       "DB_CrossCut_1_HMI".tHMR.xManualCommandEnabled := "FB_CrossCuts_1_V1_00_IDB".tHMR.xManComEn;
       "DB_CrossCut_1_HMI".tHMR.tManCmd.xManJogFwdFdbk := "FB_CrossCuts_1_V1_00_IDB".tHMR.tManCmd.xManJogFwdFdbk;
       "DB_CrossCut_1_HMI".tHMR.tManCmd.xManJogBckFdbk := "FB_CrossCuts_1_V1_00_IDB".tHMR.tManCmd.xManJogBckFdbk;
       "DB_CrossCut_1_HMI".tHMR.tManCmd.xManCarriageDownFdbk := "FB_CrossCuts_1_V1_00_IDB".tHMR.tManCmd.xManCarriageDownFdbk;
       "DB_CrossCut_1_HMI".tHMR.tManCmd.xManFireONFdbk := "FB_CrossCuts_1_V1_00_IDB".tHMR.tManCmd.xManFireONFdbk;
       "DB_CrossCut_1_HMI".tHMR.tManCmd.xManOilONFdbk := "FB_CrossCuts_1_V1_00_IDB".tHMR.tManCmd.xManOilONFdbk;

       "DB_CrossCut_1_HMI".tHMR.dDistanceSnaproll_cmm := "FB_CrossCuts_1_V1_00_IDB".tHMR.dDistanceFromSnaproll_cmm;
       "DB_CrossCut_1_HMI".tHMR.dStatus := "FB_CrossCuts_1_V1_00_IDB".tHMR.dStatus;
       "DB_CrossCut_1_HMI".tHMR.dXCutActualStatus := "FB_CrossCuts_1_V1_00_IDB".tHMR.dXCutActualStatus;
       "DB_CrossCut_1_HMI".tHMR.dXCutStatusRequest:="FB_CrossCuts_1_V1_00_IDB".tHMR.dXCutStatusRequest;
       "DB_CrossCut_1_HMI".tHMR.dDistanceFromCenterLine_cmm := "FB_CrossCuts_1_V1_00_IDB".tHMR.dDistanceFromCenterLine_cmm;
       "DB_CrossCut_1_HMI".tHMR.dAngleValue_uDegree := "FB_CrossCuts_1_V1_00_IDB".tHMR.dAngleValue_uDegree;
       "DB_CrossCut_1_HMI".tHMR.dActualCutPosRequest := "FB_CrossCuts_1_V1_00_IDB".tHMR.dActualCutPosRequest;
       "DB_CrossCut_1_HMI".tHMR.dCarriagePosition_cmm := "FB_CrossCuts_1_V1_00_IDB".tHMR.dCarriagePosition_cmm;

       "DB_CrossCut_1_HMI".tHMR.rHeadUsage_km := "FB_CrossCuts_1_V1_00_IDB".tHMR.rHeadUsage_km;

       //Move CROSS CUT #1 HMW 
       "FB_CrossCuts_1_V1_00_IDB".tHMW.xCutBreakEnabled := "DB_CrossCut_1_HMI".tHMW.xCutBreakEnabled;
       "FB_CrossCuts_1_V1_00_IDB".tHMW.xUpdateDistSnap := "DB_CrossCut_1_HMI".tHMW.xUpdateDistanceSnaproll;
       "FB_CrossCuts_1_V1_00_IDB".tHMW.xUpdateAngleValue := "DB_CrossCut_1_HMI".tHMW.xUpdateAngleValue;
       "FB_CrossCuts_1_V1_00_IDB".tHMW.xIncAngleValue := "DB_CrossCut_1_HMI".tHMW.xIncAngleValue;
       "FB_CrossCuts_1_V1_00_IDB".tHMW.xDecAngleValue := "DB_CrossCut_1_HMI".tHMW.xDecAngleValue;
       "FB_CrossCuts_1_V1_00_IDB".tHMW.xUpdateDistCenterLine := "DB_CrossCut_1_HMI".tHMW.xUpdateDistCenterLine;
       "FB_CrossCuts_1_V1_00_IDB".tHMW.xCalibDistRequest := "DB_CrossCut_1_HMI".tHMW.xCalibDistRequest;
       "FB_CrossCuts_1_V1_00_IDB".tHMW.xCalibDiagRequest := "DB_CrossCut_1_HMI".tHMW.xCalibDiagRequest;
       "FB_CrossCuts_1_V1_00_IDB".tHMW.xCutOperator := "DB_CrossCut_1_HMI".tHMW.xCutOperator;
       "FB_CrossCuts_1_V1_00_IDB".tHMW.xCutGross := "DB_CrossCut_1_HMI".tHMW.xCutGross;
       "FB_CrossCuts_1_V1_00_IDB".tHMW.xCutNet := "DB_CrossCut_1_HMI".tHMW.xCutNet;
       "FB_CrossCuts_1_V1_00_IDB".tHMW.xCutYCut := "DB_CrossCut_1_HMI".tHMW.xCutYCut;
       "FB_CrossCuts_1_V1_00_IDB".tHMW.xEnDisManCom := "DB_CrossCut_1_HMI".tHMW.xEnableManualCommand;
       "FB_CrossCuts_1_V1_00_IDB".tHMW.xResetHeadUsage := "DB_CrossCut_1_HMI".tHMW.xResetHeadUsage;

       "FB_CrossCuts_1_V1_00_IDB".tHMW.tManCmd.xMan_JogForward := "DB_CrossCut_1_HMI".tHMW.tManCmd.xMan_JogForward;
       "FB_CrossCuts_1_V1_00_IDB".tHMW.tManCmd.xMan_JobBackward := "DB_CrossCut_1_HMI".tHMW.tManCmd.xMan_JobBackward;
       "FB_CrossCuts_1_V1_00_IDB".tHMW.tManCmd.xMan_CarriageDown := "DB_CrossCut_1_HMI".tHMW.tManCmd.xMan_CarriageDown;
       "FB_CrossCuts_1_V1_00_IDB".tHMW.tManCmd.xMan_FireOn := "DB_CrossCut_1_HMI".tHMW.tManCmd.xMan_FireOn;
       "FB_CrossCuts_1_V1_00_IDB".tHMW.tManCmd.xMan_OilOn := "DB_CrossCut_1_HMI".tHMW.tManCmd.xMan_OilOn;



      "FB_CrossCuts_1_V1_00_IDB".tHMW.dOperStartCutPos_cmm := "DB_CrossCut_1_HMI".tHMW.dOperStartCutPos_cmm;
      "FB_CrossCuts_1_V1_00_IDB".tHMW.dOperEndCutPos_cmm := "DB_CrossCut_1_HMI".tHMW.dOperEndCutPos_cmm;
      "FB_CrossCuts_1_V1_00_IDB".tHMW.dDescReactTime_ms := "DB_CrossCut_1_HMI".tHMW.dDescReactTime_ms;
      "FB_CrossCuts_1_V1_00_IDB".tHMW.dRaiseReactTime_ms := "DB_CrossCut_1_HMI".tHMW.dRaiseReactTime_ms;

      "FB_CrossCuts_1_V1_00_IDB".tHMW.dFireONReactTime_ms := "DB_CrossCut_1_HMI".tHMW.dFireONReactTime_ms;
      "FB_CrossCuts_1_V1_00_IDB".tHMW.dFireOFFReactTime_ms := "DB_CrossCut_1_HMI".tHMW.dFireOFFReactTime_ms;
      "FB_CrossCuts_1_V1_00_IDB".tHMW.dOilONDelay_ms := "DB_CrossCut_1_HMI".tHMW.dOilONDelay_ms;
      "FB_CrossCuts_1_V1_00_IDB".tHMW.dOilOFFDelay_ms := "DB_CrossCut_1_HMI".tHMW.dOilOFFDelay_ms;

      "FB_CrossCuts_1_V1_00_IDB".tHMW.dCutStartOffsetDelay_cmm := "DB_CrossCut_1_HMI".tHMW.dCutStartOffsetDelay_cmm;
      "FB_CrossCuts_1_V1_00_IDB".tHMW.dCutEndOffsetDelay_cmm := "DB_CrossCut_1_HMI".tHMW.dCutEndOffsetDelay_cmm;

      "FB_CrossCuts_1_V1_00_IDB".tHMW.dDistanceFromSnaproll_cmm := "DB_CrossCut_1_HMI".tHMW.dDistanceSnaproll_cmm;
      "FB_CrossCuts_1_V1_00_IDB".tHMW.dAngleValue_uDegree := "DB_CrossCut_1_HMI".tHMW.dAngleValue_uDegree;
      "FB_CrossCuts_1_V1_00_IDB".tHMW.dDistanceFromCenterLine_cmm := "DB_CrossCut_1_HMI".tHMW.dDistanceFromCenterLine_cmm;
      "FB_CrossCuts_1_V1_00_IDB".tHMW.dDistTeoLength_cmm := "DB_CrossCut_1_HMI".tHMW.dDistTeoLength_cmm;
      "FB_CrossCuts_1_V1_00_IDB".tHMW.dDistRealLength_cmm := "DB_CrossCut_1_HMI".tHMW.dDistRealLength_cmm;

      "FB_CrossCuts_1_V1_00_IDB".tHMW.dDiagRealWidth_cmm := "DB_CrossCut_1_HMI".tHMW.dDiagRealWidth_cmm;
       "FB_CrossCuts_1_V1_00_IDB".tHMW.dDiagRealLength_cmm := "DB_CrossCut_1_HMI".tHMW.dDiagRealLength_cmm;
       "FB_CrossCuts_1_V1_00_IDB".tHMW.dDiagGlassFlow_cmm := "DB_CrossCut_1_HMI".tHMW.dDiagGlassFlow_cmm;
       "FB_CrossCuts_1_V1_00_IDB".tHMW.dDiagGlassOppFlow_cmm := "DB_CrossCut_1_HMI".tHMW.dDiagGlassOppFlow_cmm;

       "FB_CrossCuts_1_V1_00_IDB".tHMW.dCuttingPressure_mN := "DB_CrossCut_1_HMI".tHMW.dCuttingPressure_mN;
       "FB_CrossCuts_1_V1_00_IDB".tHMW.dPosOffset_cmm := "DB_CrossCut_1_HMI".tHMW.dPosOffset_cmm;

       "FB_CrossCuts_1_V1_00_IDB".tHMW.dCutPriority := "DB_CrossCut_1_HMI".tHMW.dCutPriority;

       //Move CROSS CUT #1 ALM
       "DB_CrossCut_1_HMI".tALM := "FB_CrossCuts_1_V1_00_IDB".tALM;



       //Move CROSS CUT #2 HMR 

       "DB_CrossCut_2_HMI".tHMR.xManualCommandEnabled := "FB_CrossCuts_2_V1_00_IDB".tHMR.xManComEn;
       "DB_CrossCut_2_HMI".tHMR.tManCmd.xManJogFwdFdbk := "FB_CrossCuts_2_V1_00_IDB".tHMR.tManCmd.xManJogFwdFdbk;
       "DB_CrossCut_2_HMI".tHMR.tManCmd.xManJogBckFdbk := "FB_CrossCuts_2_V1_00_IDB".tHMR.tManCmd.xManJogBckFdbk;
       "DB_CrossCut_2_HMI".tHMR.tManCmd.xManCarriageDownFdbk := "FB_CrossCuts_2_V1_00_IDB".tHMR.tManCmd.xManCarriageDownFdbk;
       "DB_CrossCut_2_HMI".tHMR.tManCmd.xManFireONFdbk := "FB_CrossCuts_2_V1_00_IDB".tHMR.tManCmd.xManFireONFdbk;
       "DB_CrossCut_2_HMI".tHMR.tManCmd.xManOilONFdbk := "FB_CrossCuts_2_V1_00_IDB".tHMR.tManCmd.xManOilONFdbk;

       "DB_CrossCut_2_HMI".tHMR.dDistanceSnaproll_cmm := "FB_CrossCuts_2_V1_00_IDB".tHMR.dDistanceFromSnaproll_cmm;
       "DB_CrossCut_2_HMI".tHMR.dStatus := "FB_CrossCuts_2_V1_00_IDB".tHMR.dStatus;
       "DB_CrossCut_2_HMI".tHMR.dXCutActualStatus := "FB_CrossCuts_2_V1_00_IDB".tHMR.dXCutActualStatus;
       "DB_CrossCut_2_HMI".tHMR.dXCutStatusRequest := "FB_CrossCuts_2_V1_00_IDB".tHMR.dXCutStatusRequest;
       "DB_CrossCut_2_HMI".tHMR.dDistanceFromCenterLine_cmm := "FB_CrossCuts_2_V1_00_IDB".tHMR.dDistanceFromCenterLine_cmm;
       "DB_CrossCut_2_HMI".tHMR.dAngleValue_uDegree := "FB_CrossCuts_2_V1_00_IDB".tHMR.dAngleValue_uDegree;
       "DB_CrossCut_2_HMI".tHMR.dActualCutPosRequest := "FB_CrossCuts_2_V1_00_IDB".tHMR.dActualCutPosRequest;
       "DB_CrossCut_2_HMI".tHMR.dCarriagePosition_cmm := "FB_CrossCuts_2_V1_00_IDB".tHMR.dCarriagePosition_cmm;

       "DB_CrossCut_2_HMI".tHMR.rHeadUsage_km := "FB_CrossCuts_2_V1_00_IDB".tHMR.rHeadUsage_km;

       //Move CROSS CUT #2 HMW 
       "FB_CrossCuts_2_V1_00_IDB".tHMW.xCutBreakEnabled := "DB_CrossCut_2_HMI".tHMW.xCutBreakEnabled;
       "FB_CrossCuts_2_V1_00_IDB".tHMW.xUpdateDistSnap := "DB_CrossCut_2_HMI".tHMW.xUpdateDistanceSnaproll;
       "FB_CrossCuts_2_V1_00_IDB".tHMW.xUpdateAngleValue := "DB_CrossCut_2_HMI".tHMW.xUpdateAngleValue;
       "FB_CrossCuts_2_V1_00_IDB".tHMW.xIncAngleValue := "DB_CrossCut_2_HMI".tHMW.xIncAngleValue;
       "FB_CrossCuts_2_V1_00_IDB".tHMW.xDecAngleValue := "DB_CrossCut_2_HMI".tHMW.xDecAngleValue;
       "FB_CrossCuts_2_V1_00_IDB".tHMW.xUpdateDistCenterLine := "DB_CrossCut_2_HMI".tHMW.xUpdateDistCenterLine;
       "FB_CrossCuts_2_V1_00_IDB".tHMW.xCalibDistRequest := "DB_CrossCut_2_HMI".tHMW.xCalibDistRequest;
       "FB_CrossCuts_2_V1_00_IDB".tHMW.xCalibDiagRequest := "DB_CrossCut_2_HMI".tHMW.xCalibDiagRequest;
       "FB_CrossCuts_2_V1_00_IDB".tHMW.xCutOperator := "DB_CrossCut_2_HMI".tHMW.xCutOperator;
       "FB_CrossCuts_2_V1_00_IDB".tHMW.xCutGross := "DB_CrossCut_2_HMI".tHMW.xCutGross;
       "FB_CrossCuts_2_V1_00_IDB".tHMW.xCutNet := "DB_CrossCut_2_HMI".tHMW.xCutNet;
       "FB_CrossCuts_2_V1_00_IDB".tHMW.xCutYCut := "DB_CrossCut_2_HMI".tHMW.xCutYCut;
       "FB_CrossCuts_2_V1_00_IDB".tHMW.xEnDisManCom := "DB_CrossCut_2_HMI".tHMW.xEnableManualCommand;
       "FB_CrossCuts_2_V1_00_IDB".tHMW.xResetHeadUsage := "DB_CrossCut_2_HMI".tHMW.xResetHeadUsage;

       "FB_CrossCuts_2_V1_00_IDB".tHMW.tManCmd.xMan_JogForward := "DB_CrossCut_2_HMI".tHMW.tManCmd.xMan_JogForward;
       "FB_CrossCuts_2_V1_00_IDB".tHMW.tManCmd.xMan_JobBackward := "DB_CrossCut_2_HMI".tHMW.tManCmd.xMan_JobBackward;
       "FB_CrossCuts_2_V1_00_IDB".tHMW.tManCmd.xMan_CarriageDown := "DB_CrossCut_2_HMI".tHMW.tManCmd.xMan_CarriageDown;
       "FB_CrossCuts_2_V1_00_IDB".tHMW.tManCmd.xMan_FireOn := "DB_CrossCut_2_HMI".tHMW.tManCmd.xMan_FireOn;
       "FB_CrossCuts_2_V1_00_IDB".tHMW.tManCmd.xMan_OilOn := "DB_CrossCut_2_HMI".tHMW.tManCmd.xMan_OilOn;



       "FB_CrossCuts_2_V1_00_IDB".tHMW.dOperStartCutPos_cmm := "DB_CrossCut_2_HMI".tHMW.dOperStartCutPos_cmm;
       "FB_CrossCuts_2_V1_00_IDB".tHMW.dOperEndCutPos_cmm := "DB_CrossCut_2_HMI".tHMW.dOperEndCutPos_cmm;
       "FB_CrossCuts_2_V1_00_IDB".tHMW.dDescReactTime_ms := "DB_CrossCut_2_HMI".tHMW.dDescReactTime_ms;
       "FB_CrossCuts_2_V1_00_IDB".tHMW.dRaiseReactTime_ms := "DB_CrossCut_2_HMI".tHMW.dRaiseReactTime_ms;

       "FB_CrossCuts_2_V1_00_IDB".tHMW.dFireONReactTime_ms := "DB_CrossCut_2_HMI".tHMW.dFireONReactTime_ms;
       "FB_CrossCuts_2_V1_00_IDB".tHMW.dFireOFFReactTime_ms := "DB_CrossCut_2_HMI".tHMW.dFireOFFReactTime_ms;
       "FB_CrossCuts_2_V1_00_IDB".tHMW.dOilONDelay_ms := "DB_CrossCut_2_HMI".tHMW.dOilONDelay_ms;
       "FB_CrossCuts_2_V1_00_IDB".tHMW.dOilOFFDelay_ms := "DB_CrossCut_2_HMI".tHMW.dOilOFFDelay_ms;

       "FB_CrossCuts_2_V1_00_IDB".tHMW.dCutStartOffsetDelay_cmm := "DB_CrossCut_2_HMI".tHMW.dCutStartOffsetDelay_cmm;
       "FB_CrossCuts_2_V1_00_IDB".tHMW.dCutEndOffsetDelay_cmm := "DB_CrossCut_2_HMI".tHMW.dCutEndOffsetDelay_cmm;

       "FB_CrossCuts_2_V1_00_IDB".tHMW.dDistanceFromSnaproll_cmm := "DB_CrossCut_2_HMI".tHMW.dDistanceSnaproll_cmm;
       "FB_CrossCuts_2_V1_00_IDB".tHMW.dAngleValue_uDegree := "DB_CrossCut_2_HMI".tHMW.dAngleValue_uDegree;
       "FB_CrossCuts_2_V1_00_IDB".tHMW.dDistanceFromCenterLine_cmm := "DB_CrossCut_2_HMI".tHMW.dDistanceFromCenterLine_cmm;
       "FB_CrossCuts_2_V1_00_IDB".tHMW.dDistTeoLength_cmm := "DB_CrossCut_2_HMI".tHMW.dDistTeoLength_cmm;
       "FB_CrossCuts_2_V1_00_IDB".tHMW.dDistRealLength_cmm := "DB_CrossCut_2_HMI".tHMW.dDistRealLength_cmm;

       "FB_CrossCuts_2_V1_00_IDB".tHMW.dDiagRealWidth_cmm := "DB_CrossCut_2_HMI".tHMW.dDiagRealWidth_cmm;
       "FB_CrossCuts_2_V1_00_IDB".tHMW.dDiagRealLength_cmm := "DB_CrossCut_2_HMI".tHMW.dDiagRealLength_cmm;
       "FB_CrossCuts_2_V1_00_IDB".tHMW.dDiagGlassFlow_cmm := "DB_CrossCut_2_HMI".tHMW.dDiagGlassFlow_cmm;
       "FB_CrossCuts_2_V1_00_IDB".tHMW.dDiagGlassOppFlow_cmm := "DB_CrossCut_2_HMI".tHMW.dDiagGlassOppFlow_cmm;

       "FB_CrossCuts_2_V1_00_IDB".tHMW.dCuttingPressure_mN := "DB_CrossCut_2_HMI".tHMW.dCuttingPressure_mN;
       "FB_CrossCuts_2_V1_00_IDB".tHMW.dPosOffset_cmm := "DB_CrossCut_2_HMI".tHMW.dPosOffset_cmm;

       "FB_CrossCuts_2_V1_00_IDB".tHMW.dCutPriority := "DB_CrossCut_2_HMI".tHMW.dCutPriority;

       //Move CROSS CUT #2 ALM
       "DB_CrossCut_2_HMI".tALM := "FB_CrossCuts_2_V1_00_IDB".tALM;



       //Move CROSS CUT #3 HMR 

       "DB_CrossCut_3_HMI".tHMR.xManualCommandEnabled := "FB_CrossCuts_3_V1_00_IDB".tHMR.xManComEn;
       "DB_CrossCut_3_HMI".tHMR.tManCmd.xManJogFwdFdbk := "FB_CrossCuts_3_V1_00_IDB".tHMR.tManCmd.xManJogFwdFdbk;
       "DB_CrossCut_3_HMI".tHMR.tManCmd.xManJogBckFdbk := "FB_CrossCuts_3_V1_00_IDB".tHMR.tManCmd.xManJogBckFdbk;
       "DB_CrossCut_3_HMI".tHMR.tManCmd.xManCarriageDownFdbk := "FB_CrossCuts_3_V1_00_IDB".tHMR.tManCmd.xManCarriageDownFdbk;
       "DB_CrossCut_3_HMI".tHMR.tManCmd.xManFireONFdbk := "FB_CrossCuts_3_V1_00_IDB".tHMR.tManCmd.xManFireONFdbk;
       "DB_CrossCut_3_HMI".tHMR.tManCmd.xManOilONFdbk := "FB_CrossCuts_3_V1_00_IDB".tHMR.tManCmd.xManOilONFdbk;

       "DB_CrossCut_3_HMI".tHMR.dDistanceSnaproll_cmm := "FB_CrossCuts_3_V1_00_IDB".tHMR.dDistanceFromSnaproll_cmm;
       "DB_CrossCut_3_HMI".tHMR.dStatus := "FB_CrossCuts_3_V1_00_IDB".tHMR.dStatus;
       "DB_CrossCut_3_HMI".tHMR.dXCutActualStatus := "FB_CrossCuts_3_V1_00_IDB".tHMR.dXCutActualStatus;
       "DB_CrossCut_3_HMI".tHMR.dXCutStatusRequest := "FB_CrossCuts_3_V1_00_IDB".tHMR.dXCutStatusRequest;
       "DB_CrossCut_3_HMI".tHMR.dDistanceFromCenterLine_cmm := "FB_CrossCuts_3_V1_00_IDB".tHMR.dDistanceFromCenterLine_cmm;
       "DB_CrossCut_3_HMI".tHMR.dAngleValue_uDegree := "FB_CrossCuts_3_V1_00_IDB".tHMR.dAngleValue_uDegree;
       "DB_CrossCut_3_HMI".tHMR.dActualCutPosRequest := "FB_CrossCuts_3_V1_00_IDB".tHMR.dActualCutPosRequest;
       "DB_CrossCut_3_HMI".tHMR.dCarriagePosition_cmm := "FB_CrossCuts_3_V1_00_IDB".tHMR.dCarriagePosition_cmm;

       "DB_CrossCut_3_HMI".tHMR.rHeadUsage_km := "FB_CrossCuts_3_V1_00_IDB".tHMR.rHeadUsage_km;

       //Move CROSS CUT #3 HMW 
       "FB_CrossCuts_3_V1_00_IDB".tHMW.xCutBreakEnabled := "DB_CrossCut_3_HMI".tHMW.xCutBreakEnabled;
       "FB_CrossCuts_3_V1_00_IDB".tHMW.xUpdateDistSnap := "DB_CrossCut_3_HMI".tHMW.xUpdateDistanceSnaproll;
       "FB_CrossCuts_3_V1_00_IDB".tHMW.xUpdateAngleValue := "DB_CrossCut_3_HMI".tHMW.xUpdateAngleValue;
       "FB_CrossCuts_3_V1_00_IDB".tHMW.xIncAngleValue := "DB_CrossCut_3_HMI".tHMW.xIncAngleValue;
       "FB_CrossCuts_3_V1_00_IDB".tHMW.xDecAngleValue := "DB_CrossCut_3_HMI".tHMW.xDecAngleValue;
       "FB_CrossCuts_3_V1_00_IDB".tHMW.xUpdateDistCenterLine := "DB_CrossCut_3_HMI".tHMW.xUpdateDistCenterLine;
       "FB_CrossCuts_3_V1_00_IDB".tHMW.xCalibDistRequest := "DB_CrossCut_3_HMI".tHMW.xCalibDistRequest;
       "FB_CrossCuts_3_V1_00_IDB".tHMW.xCalibDiagRequest := "DB_CrossCut_3_HMI".tHMW.xCalibDiagRequest;
       "FB_CrossCuts_3_V1_00_IDB".tHMW.xCutOperator := "DB_CrossCut_3_HMI".tHMW.xCutOperator;
       "FB_CrossCuts_3_V1_00_IDB".tHMW.xCutGross := "DB_CrossCut_3_HMI".tHMW.xCutGross;
       "FB_CrossCuts_3_V1_00_IDB".tHMW.xCutNet := "DB_CrossCut_3_HMI".tHMW.xCutNet;
       "FB_CrossCuts_3_V1_00_IDB".tHMW.xCutYCut := "DB_CrossCut_3_HMI".tHMW.xCutYCut;
       "FB_CrossCuts_3_V1_00_IDB".tHMW.xEnDisManCom := "DB_CrossCut_3_HMI".tHMW.xEnableManualCommand;
       "FB_CrossCuts_3_V1_00_IDB".tHMW.xResetHeadUsage := "DB_CrossCut_3_HMI".tHMW.xResetHeadUsage;

       "FB_CrossCuts_3_V1_00_IDB".tHMW.tManCmd.xMan_JogForward := "DB_CrossCut_3_HMI".tHMW.tManCmd.xMan_JogForward;
       "FB_CrossCuts_3_V1_00_IDB".tHMW.tManCmd.xMan_JobBackward := "DB_CrossCut_3_HMI".tHMW.tManCmd.xMan_JobBackward;
       "FB_CrossCuts_3_V1_00_IDB".tHMW.tManCmd.xMan_CarriageDown := "DB_CrossCut_3_HMI".tHMW.tManCmd.xMan_CarriageDown;
       "FB_CrossCuts_3_V1_00_IDB".tHMW.tManCmd.xMan_FireOn := "DB_CrossCut_3_HMI".tHMW.tManCmd.xMan_FireOn;
       "FB_CrossCuts_3_V1_00_IDB".tHMW.tManCmd.xMan_OilOn := "DB_CrossCut_3_HMI".tHMW.tManCmd.xMan_OilOn;



       "FB_CrossCuts_3_V1_00_IDB".tHMW.dOperStartCutPos_cmm := "DB_CrossCut_3_HMI".tHMW.dOperStartCutPos_cmm;
       "FB_CrossCuts_3_V1_00_IDB".tHMW.dOperEndCutPos_cmm := "DB_CrossCut_3_HMI".tHMW.dOperEndCutPos_cmm;
       "FB_CrossCuts_3_V1_00_IDB".tHMW.dDescReactTime_ms := "DB_CrossCut_3_HMI".tHMW.dDescReactTime_ms;
       "FB_CrossCuts_3_V1_00_IDB".tHMW.dRaiseReactTime_ms := "DB_CrossCut_3_HMI".tHMW.dRaiseReactTime_ms;

       "FB_CrossCuts_3_V1_00_IDB".tHMW.dFireONReactTime_ms := "DB_CrossCut_3_HMI".tHMW.dFireONReactTime_ms;
       "FB_CrossCuts_3_V1_00_IDB".tHMW.dFireOFFReactTime_ms := "DB_CrossCut_3_HMI".tHMW.dFireOFFReactTime_ms;
       "FB_CrossCuts_3_V1_00_IDB".tHMW.dOilONDelay_ms := "DB_CrossCut_3_HMI".tHMW.dOilONDelay_ms;
       "FB_CrossCuts_3_V1_00_IDB".tHMW.dOilOFFDelay_ms := "DB_CrossCut_3_HMI".tHMW.dOilOFFDelay_ms;

       "FB_CrossCuts_3_V1_00_IDB".tHMW.dCutStartOffsetDelay_cmm := "DB_CrossCut_3_HMI".tHMW.dCutStartOffsetDelay_cmm;
       "FB_CrossCuts_3_V1_00_IDB".tHMW.dCutEndOffsetDelay_cmm := "DB_CrossCut_3_HMI".tHMW.dCutEndOffsetDelay_cmm;

       "FB_CrossCuts_3_V1_00_IDB".tHMW.dDistanceFromSnaproll_cmm := "DB_CrossCut_3_HMI".tHMW.dDistanceSnaproll_cmm;
       "FB_CrossCuts_3_V1_00_IDB".tHMW.dAngleValue_uDegree := "DB_CrossCut_3_HMI".tHMW.dAngleValue_uDegree;
       "FB_CrossCuts_3_V1_00_IDB".tHMW.dDistanceFromCenterLine_cmm := "DB_CrossCut_3_HMI".tHMW.dDistanceFromCenterLine_cmm;
       "FB_CrossCuts_3_V1_00_IDB".tHMW.dDistTeoLength_cmm := "DB_CrossCut_3_HMI".tHMW.dDistTeoLength_cmm;
       "FB_CrossCuts_3_V1_00_IDB".tHMW.dDistRealLength_cmm := "DB_CrossCut_3_HMI".tHMW.dDistRealLength_cmm;

       "FB_CrossCuts_3_V1_00_IDB".tHMW.dDiagRealWidth_cmm := "DB_CrossCut_3_HMI".tHMW.dDiagRealWidth_cmm;
       "FB_CrossCuts_3_V1_00_IDB".tHMW.dDiagRealLength_cmm := "DB_CrossCut_3_HMI".tHMW.dDiagRealLength_cmm;
       "FB_CrossCuts_3_V1_00_IDB".tHMW.dDiagGlassFlow_cmm := "DB_CrossCut_3_HMI".tHMW.dDiagGlassFlow_cmm;
       "FB_CrossCuts_3_V1_00_IDB".tHMW.dDiagGlassOppFlow_cmm := "DB_CrossCut_3_HMI".tHMW.dDiagGlassOppFlow_cmm;

       "FB_CrossCuts_3_V1_00_IDB".tHMW.dCuttingPressure_mN := "DB_CrossCut_3_HMI".tHMW.dCuttingPressure_mN;
       "FB_CrossCuts_3_V1_00_IDB".tHMW.dPosOffset_cmm := "DB_CrossCut_3_HMI".tHMW.dPosOffset_cmm;

       "FB_CrossCuts_3_V1_00_IDB".tHMW.dCutPriority := "DB_CrossCut_3_HMI".tHMW.dCutPriority;

       //Move CROSS CUT #3 ALM
       "DB_CrossCut_3_HMI".tALM := "FB_CrossCuts_3_V1_00_IDB".tALM;



       //Move YCUT 1 HMR
       "DB_YCut_1_HMI".tHMR.dDistanceSnaproll_cmm := "FB_YCuts1_V1_00_IDB".tHMR.dDistanceFromSnaproll_cmm;
       //Move YCUT 1  HMW
       "FB_YCuts1_V1_00_IDB".tHMW.xUpdateDistSnap := "DB_YCut_1_HMI".tHMW.xUpdateDistanceSnaproll;
       "FB_YCuts1_V1_00_IDB".tHMW.dDistanceFromSnaproll_cmm := "DB_YCut_1_HMI".tHMW.dDistanceSnaproll_cmm;
       //Move YCUT 1  ALM 
       "DB_YCut_1_HMI".tALM.tF := "FB_YCuts1_V1_00_IDB".tALM.tF;
       "DB_YCut_1_HMI".tALM.tS := "FB_YCuts1_V1_00_IDB".tALM.tS;
       "DB_YCut_1_HMI".tALM.tW:= "FB_YCuts1_V1_00_IDB".tALM.tW;

       //Move YCUT 2 HMR
       "DB_YCut_2_HMI".tHMR.dDistanceSnaproll_cmm := "FB_YCuts2_V1_00_IDB".tHMR.dDistanceFromSnaproll_cmm;
       //Move YCUT 2  HMW
       "FB_YCuts2_V1_00_IDB".tHMW.xUpdateDistSnap := "DB_YCut_2_HMI".tHMW.xUpdateDistanceSnaproll;
       "FB_YCuts2_V1_00_IDB".tHMW.dDistanceFromSnaproll_cmm := "DB_YCut_2_HMI".tHMW.dDistanceSnaproll_cmm;
       //Move YCUT 1  ALM 
       "DB_YCut_2_HMI".tALM.tF := "FB_YCuts2_V1_00_IDB".tALM.tF;
       "DB_YCut_2_HMI".tALM.tS := "FB_YCuts2_V1_00_IDB".tALM.tS;
       "DB_YCut_2_HMI".tALM.tW := "FB_YCuts2_V1_00_IDB".tALM.tW;

       //Move Marker M220 HMR
       "DB_Marker_HMI".tHMR.dSpare0 :="FB_Markers_V1.00_IDB".tHMR.dSpare;
       //Move Marker M220  HMW
       "FB_Markers_V1.00_IDB".tHMW.dSpare :=  "DB_Marker_HMI".tHMW.dSpare0;
       //Move Marker M220 ALM  
       "DB_Marker_HMI".tALM.tF := "FB_Markers_V1.00_IDB".tALM.tF;
       "DB_Marker_HMI".tALM.tS := "FB_Markers_V1.00_IDB".tALM.tS;
       "DB_Marker_HMI".tALM.tW := "FB_Markers_V1.00_IDB".tALM.tW;

       //Move DIGITIZER #1 HMR
       "DB_Digitizer_1_HMI".tHMR.xManualCommandEnabled := "FB_Digitizer_1_V1_00_IDB".tHMR.xManComEn;
       "DB_Digitizer_1_HMI".tHMR.tManCmd.xMan_DescEncFdbk:= "FB_Digitizer_1_V1_00_IDB".tHMR.xMan_DescEncFdbk;
       "DB_Digitizer_1_HMI".tHMR.dEncoderStatus := "FB_Digitizer_1_V1_00_IDB".tHMR.dEncoderStatus;
       "DB_Digitizer_1_HMI".tHMR.dFm152Status := "FB_Digitizer_1_V1_00_IDB".tHMR.dFm152Status;
       "DB_Digitizer_1_HMI".tHMR.dActualEncoderSpeed_mm_min := "FB_Digitizer_1_V1_00_IDB".tHMR.dActualEncoderSpeed_mm_min;
       "DB_Digitizer_1_HMI".tHMR.dCalibrationF1Unit_unit := "FB_Digitizer_1_V1_00_IDB".tHMR.dCalibrationF1Unit_unit;
       "DB_Digitizer_1_HMI".tHMR.dCalibrationF2Unit_unit := "FB_Digitizer_1_V1_00_IDB".tHMR.dCalibrationF2Unit_unit;
       "DB_Digitizer_1_HMI".tHMR.dCalibrationCardF1Unit_unit := "FB_Digitizer_1_V1_00_IDB".tHMR.dCalibrationCardF1Unit_unit;
       "DB_Digitizer_1_HMI".tHMR.dCalibrationCardF2Unit_unit := "FB_Digitizer_1_V1_00_IDB".tHMR.dCalibrationCardF2Unit_unit;


       //Move DIGITIZER #1  HMW
       "FB_Digitizer_1_V1_00_IDB".tHMW.xCalibUpdateF1 := "DB_Digitizer_1_HMI".tHMW.xCalibRequest;
       "FB_Digitizer_1_V1_00_IDB".tHMW.xCalibUpdateF2 := "DB_Digitizer_1_HMI".tHMW.xCalibUpdateF1;
       "FB_Digitizer_1_V1_00_IDB".tHMW.xCalibRequest := "DB_Digitizer_1_HMI".tHMW.xCalibUpdateF2;
       "FB_Digitizer_1_V1_00_IDB".tHMW.xMan_DescentEnc:="DB_Digitizer_1_HMI".tHMW.tManCmd.xMan_DescentEnc;
       "FB_Digitizer_1_V1_00_IDB".tHMW.xGlassSensorEnabled := "DB_Digitizer_1_HMI".tHMW.xGlassSensorEnabled;
       "FB_Digitizer_1_V1_00_IDB".tHMW.xEnDisManCom := "DB_Digitizer_1_HMI".tHMW.xEnableManualCommand;
       "FB_Digitizer_1_V1_00_IDB".tHMW.dCalibTheoLength_cmm := "DB_Digitizer_1_HMI".tHMW.dCalibTheoLength_cmm;
       "FB_Digitizer_1_V1_00_IDB".tHMW.dCalibRealLength_cmm := "DB_Digitizer_1_HMI".tHMW.dCalibRealLength_cmm;
       "FB_Digitizer_1_V1_00_IDB".tHMW.dCalibWriteF1_unit := "DB_Digitizer_1_HMI".tHMW.dCalibWriteF1_unit;
       "FB_Digitizer_1_V1_00_IDB".tHMW.dCalibWriteF2_unit := "DB_Digitizer_1_HMI".tHMW.dCalibWriteF2_unit;
       "FB_Digitizer_1_V1_00_IDB".tHMW.dRequestJogSpeed_mm_min := "DB_Digitizer_1_HMI".tHMW.dRequestJogSpeed_mm_min;




       //Move DIGITIZER #1 ALM  
       "DB_Digitizer_1_HMI".tALM.tS := "FB_Digitizer_1_V1_00_IDB".tALM.tS;
       "DB_Digitizer_1_HMI".tALM.tF := "FB_Digitizer_1_V1_00_IDB".tALM.tF;
       "DB_Digitizer_1_HMI".tALM.tW := "FB_Digitizer_1_V1_00_IDB".tALM.tW;

       //Move DIGITIZER #2 HMR
       "DB_Digitizer_2_HMI".tHMR.xManualCommandEnabled := "FB_Digitizer_2_V1_00_IDB".tHMR.xManComEn;
       "DB_Digitizer_2_HMI".tHMR.tManCmd.xMan_DescEncFdbk := "FB_Digitizer_2_V1_00_IDB".tHMR.xMan_DescEncFdbk;
       "DB_Digitizer_2_HMI".tHMR.dEncoderStatus := "FB_Digitizer_2_V1_00_IDB".tHMR.dEncoderStatus;
       "DB_Digitizer_2_HMI".tHMR.dFm152Status := "FB_Digitizer_2_V1_00_IDB".tHMR.dFm152Status;
       "DB_Digitizer_2_HMI".tHMR.dActualEncoderSpeed_mm_min := "FB_Digitizer_2_V1_00_IDB".tHMR.dActualEncoderSpeed_mm_min;
       "DB_Digitizer_2_HMI".tHMR.dCalibrationF1Unit_unit := "FB_Digitizer_2_V1_00_IDB".tHMR.dCalibrationF1Unit_unit;
       "DB_Digitizer_2_HMI".tHMR.dCalibrationF2Unit_unit := "FB_Digitizer_2_V1_00_IDB".tHMR.dCalibrationF2Unit_unit;
       "DB_Digitizer_2_HMI".tHMR.dCalibrationCardF1Unit_unit := "FB_Digitizer_2_V1_00_IDB".tHMR.dCalibrationCardF1Unit_unit;
       "DB_Digitizer_2_HMI".tHMR.dCalibrationCardF2Unit_unit := "FB_Digitizer_2_V1_00_IDB".tHMR.dCalibrationCardF2Unit_unit;


       //Move DIGITIZER #2  HMW
       "FB_Digitizer_2_V1_00_IDB".tHMW.xCalibUpdateF1 := "DB_Digitizer_2_HMI".tHMW.xCalibRequest;
       "FB_Digitizer_2_V1_00_IDB".tHMW.xCalibUpdateF2 := "DB_Digitizer_2_HMI".tHMW.xCalibUpdateF1;
       "FB_Digitizer_2_V1_00_IDB".tHMW.xCalibRequest := "DB_Digitizer_2_HMI".tHMW.xCalibUpdateF2;
       "FB_Digitizer_2_V1_00_IDB".tHMW.xMan_DescentEnc := "DB_Digitizer_2_HMI".tHMW.tManCmd.xMan_DescentEnc;
       "FB_Digitizer_2_V1_00_IDB".tHMW.xGlassSensorEnabled := "DB_Digitizer_2_HMI".tHMW.xGlassSensorEnabled;
       "FB_Digitizer_2_V1_00_IDB".tHMW.xEnDisManCom := "DB_Digitizer_2_HMI".tHMW.xEnableManualCommand;
       "FB_Digitizer_2_V1_00_IDB".tHMW.dCalibTheoLength_cmm := "DB_Digitizer_2_HMI".tHMW.dCalibTheoLength_cmm;
       "FB_Digitizer_2_V1_00_IDB".tHMW.dCalibRealLength_cmm := "DB_Digitizer_2_HMI".tHMW.dCalibRealLength_cmm;
       "FB_Digitizer_2_V1_00_IDB".tHMW.dCalibWriteF1_unit := "DB_Digitizer_2_HMI".tHMW.dCalibWriteF1_unit;
       "FB_Digitizer_2_V1_00_IDB".tHMW.dCalibWriteF2_unit := "DB_Digitizer_2_HMI".tHMW.dCalibWriteF2_unit;
       "FB_Digitizer_2_V1_00_IDB".tHMW.dRequestJogSpeed_mm_min := "DB_Digitizer_2_HMI".tHMW.dRequestJogSpeed_mm_min;




       //Move DIGITIZER #2 ALM  
       "DB_Digitizer_2_HMI".tALM.tS := "FB_Digitizer_2_V1_00_IDB".tALM.tS;
       "DB_Digitizer_2_HMI".tALM.tF := "FB_Digitizer_2_V1_00_IDB".tALM.tF;
       "DB_Digitizer_2_HMI".tALM.tW := "FB_Digitizer_2_V1_00_IDB".tALM.tW;

       /////////////////////////////////////////////////////////////////////////////////////////////////////////



       //Move Digitizer  ALM 
       "DB_TrackENC_HMI".tALM.tS := "FB_TrackEncoder_V1_00_IDB".tALM.tS;
       "DB_TrackENC_HMI".tALM .tF :="FB_TrackEncoder_V1_00_IDB".tALM.tF;
       "DB_TrackENC_HMI".tALM.tW := "FB_TrackEncoder_V1_00_IDB".tALM.tW ;
END_FUNCTION

// folder: Library_LGF

FUNCTION "GP_GetArraySize" : Int   // FC2, SCL
TITLE = GP_GetArraySize
{ S7_Optimized_Access := 'TRUE' }
AUTHOR : Cigliutt
FAMILY : GP
VERSION : 1.0
// This FC will return the number of element of one array
   VAR_IN_OUT
      INO_vArray : Variant;   // Array to check the number of elements
   END_VAR
   VAR_TEMP
      TMP_udNumEl : UDInt;
   END_VAR
   // Ret_Val : Number of elements found. 0 if is not an array
BEGIN
   #TMP_udNumEl := 0;

   IF IS_ARRAY(#INO_vArray) THEN
       #TMP_udNumEl := CountOfElements(#INO_vArray);
   END_IF;

   #GP_GetArraySize := UDINT_TO_INT(#TMP_udNumEl);
END_FUNCTION

FUNCTION "GP_BlockMoveStruct" : Int   // FC16, SCL
TITLE = GP_BlockMoveStruct
{ S7_Optimized_Access := 'TRUE' }
AUTHOR : Cigliutt
FAMILY : GP
VERSION : 1.0
// This FC will be move data from one array of structure to another array of structure.
   VAR_INPUT
      IN_iSourceIndex : Int;   // Array source index
      IN_iDestIndex : Int;   // Array destination index
      IN_iCount : Int;   // Numer of element to move
   END_VAR
   VAR_IN_OUT
      INO_vSourceArrayStruct : Variant;   // Source array of struct
      INO_vDestArrayStruct : Variant;   // Destination array of struct
   END_VAR
   // Ret_Val : MOVE_BLK_VARIANT return
BEGIN
   #GP_BlockMoveStruct :=  MOVE_BLK_VARIANT(SRC:=#INO_vSourceArrayStruct,
                                            COUNT:=INT_TO_UDINT(#IN_iCount),
                                            SRC_INDEX:=INT_TO_DINT(#IN_iSourceIndex),
                                            DEST_INDEX:=INT_TO_DINT(#IN_iDestIndex),
                                            DEST=>#INO_vDestArrayStruct);
END_FUNCTION

FUNCTION "GP_tmONOFF_V1.00" : Void   // FC23, SCL
TITLE = Timer ON OFF
{ S7_Optimized_Access := 'TRUE' }
AUTHOR : A.Cigliutti
FAMILY : Bottero
VERSION : 1.0
   VAR_INPUT
      IN_xValue : Bool;   // Signal input
      IN_dDelayON_ms : DInt;   // Delay ON signal [ms]
      IN_dRetainOFF_ms : DInt;   // Retain OFF signal [ms]
   END_VAR
   VAR_IN_OUT
      INO_tInstance : "UDT_IECTONTOFF_V1.00";   // Bottero IEC Timer
      INO_tOBInit : "GP_OB_Initialize";   // OB Counters cicle
   END_VAR
BEGIN
   IF #IN_xValue AND NOT #INO_tInstance.INTERNAL_xLastSignalState THEN
       #INO_tInstance.INTERNAL_dWaitingON_ms := #IN_dDelayON_ms;
   ELSIF NOT #IN_xValue AND #INO_tInstance.INTERNAL_xLastSignalState THEN
       #INO_tInstance.INTERNAL_dRetainOFF_ms := #IN_dRetainOFF_ms;
   ELSIF #INO_tInstance.INTERNAL_dWaitingON_ms > 0 OR #INO_tInstance.INTERNAL_dRetainOFF_ms > 0 THEN 
       #INO_tInstance.INTERNAL_dWaitingON_ms -= #INO_tOBInit.OUT_dExecutionTime_ms;
       #INO_tInstance.INTERNAL_dRetainOFF_ms -= #INO_tOBInit.OUT_dExecutionTime_ms;
   END_IF;

   #INO_tInstance.INTERNAL_xLastSignalState := #IN_xValue;

   IF (#IN_xValue AND #INO_tInstance.INTERNAL_dWaitingON_ms <= 0) OR
       (#INO_tInstance.INTERNAL_dRetainOFF_ms > 0)  THEN
       ENO := TRUE;
       #INO_tInstance.OUT_xDone := TRUE;
   ELSE
       ENO := FALSE;
       #INO_tInstance.OUT_xDone := FALSE;
   END_IF;
END_FUNCTION

FUNCTION "GP_tmOFF_V1.00" : Void   // FC24, SCL
TITLE = Timer OFF
{ S7_Optimized_Access := 'TRUE' }
AUTHOR : A.Cigliutti
FAMILY : Bottero
VERSION : 1.0
   VAR_INPUT
      IN_xValue : Bool;   // Signal input
      IN_dRetainOFF_ms : DInt;   // Retain OFF signal [ms]
   END_VAR
   VAR_IN_OUT
      INO_tInstance : "UDT_IECTOFF_V1.00";   // Bottero IEC Timer
      INO_tOBInit : "GP_OB_Initialize";   // OB Counters cicle
   END_VAR
BEGIN
   IF NOT #IN_xValue AND #INO_tInstance.INTERNAL_xLastSignalState THEN
       #INO_tInstance.INTERNAL_dRetainOFF_ms := #IN_dRetainOFF_ms;
   ELSIF (#INO_tInstance.INTERNAL_dRetainOFF_ms > 0) THEN
       #INO_tInstance.INTERNAL_dRetainOFF_ms -= #INO_tOBInit.OUT_dExecutionTime_ms;
   END_IF;

   #INO_tInstance.INTERNAL_xLastSignalState := #IN_xValue;

   IF (#IN_xValue OR #INO_tInstance.INTERNAL_dRetainOFF_ms > 0) THEN
       ENO := TRUE;
       #INO_tInstance.OUT_xDone := TRUE;
   ELSE
       ENO := FALSE;
       #INO_tInstance.OUT_xDone := FALSE;
   END_IF;
END_FUNCTION

FUNCTION "GP_tmON_V1.00" : Void   // FC25, SCL
TITLE = Timer ON
{ S7_Optimized_Access := 'TRUE' }
AUTHOR : A.Cigliutti
FAMILY : Bottero
VERSION : 1.0
   VAR_INPUT
      IN_xValue : Bool;   // Signal input
      IN_dDelayON_ms : DInt;   // Delay ON signal [ms]
   END_VAR
   VAR_IN_OUT
      INO_tInstance : "UDT_IECTON_V1.00";   // Bottero IEC Timer
      INO_tOBInit : "GP_OB_Initialize";   // OB Counters cicle
   END_VAR
BEGIN
   IF #IN_xValue AND NOT #INO_tInstance.INTERNAL_xLastSignalState THEN
       #INO_tInstance.INTERNAL_dWaitingON_ms := #IN_dDelayON_ms;
   ELSIF (#INO_tInstance.INTERNAL_dWaitingON_ms > 0) THEN
       #INO_tInstance.INTERNAL_dWaitingON_ms-= #INO_tOBInit.OUT_dExecutionTime_ms;
   END_IF;

   #INO_tInstance.INTERNAL_xLastSignalState := #IN_xValue;

   IF (#IN_xValue AND #INO_tInstance.INTERNAL_dWaitingON_ms <= 0) THEN
       ENO := TRUE;
       #INO_tInstance.OUT_xDone := TRUE;
   ELSE
       ENO := FALSE;
       #INO_tInstance.OUT_xDone := FALSE;
   END_IF;
END_FUNCTION

// folder: Library_LGF/4 Math operations

FUNCTION "LGF_RandomRange_Dint" : DInt   // FC10013, SCL
TITLE = LGF_RandomRange_DInt
{ S7_Optimized_Access := 'TRUE' }
AUTHOR : Siemens_Digital_Industries
FAMILY : LGF
NAME : LGF_RandomRange_DInt
// This function generates random numbers in defined limits (Datatype DInt)
   VAR_INPUT
      minValue : DInt;   // minimal Value random can reach / Minimum value of the range of the random number
      maxValue : DInt;   // maximal Value random can reach / Maximum value of the range of the random number
   END_VAR
   VAR_OUTPUT
      error : Bool;   // Error if true
      status : Word;   // Status of the function
      subfunctionStatus : Word;   // Status or return value of called FB's, FCs and system blocks
   END_VAR
   VAR_TEMP
      tempTime : DTL;   // System time
      tempNanoSecondInDWord : DWord;   // UDINT converted to DWORD for access to individual bytes
      tempTimeStatus : Word;   // Status of the instruction RD_SYS_T
      tempRandomValue : DWord;   // Random-start-value
      tempNormReal : Real;   // Normalized value
   END_VAR
   // Ret_Val : Returns random DInt number in a predefined range
   VAR CONSTANT
      ZERO : DInt := 0;   // Zero value in case of error
      MAX_UDINT : UDInt := 4294967295 ;   // Maximum UDINT value
      SUB_STATUS_NO_ERROR : Word := 16#0000;   // Status: sub function call ends without error
      STATUS_FINISHED_NO_ERROR : Word := 16#0000;   // Status: Execution finished without errors
      ERR_MAX_LESS_MIN : Word := 16#8200;   // Error: The maximum limit number is smaller than the minimum limit number
      ERR_RD_SYS_T : Word := 16#8600;   // Error: System function Read system time returned an error
   END_VAR
BEGIN
   REGION Block info header
     //=============================================================================
     // SIEMENS AG / (c)Copyright 2017
     //-----------------------------------------------------------------------------
     // Title:            LGF_RandomRange_DInt
     // Comment/Function: This function generates random numbers in defined limits (Datatype DInt)
     // Library/Family:   LGF(Library General Functions)
     // Author:           Siemens Digital Industry Support
     // Tested with:      S7-PLCSIM Advanced V2.0 SP1
     // Engineering:      TIA Portal V15 Update 2
     // Restrictions:     ENO disabled - error handling done by error and status
     // Requirements:     PLC (S7-1200 / S7-1500)
     //-------------------------------------------------------------------------------
     // Change log table:
     // Version  | Date       | Expert in charge       | Changes applied
     //----------|------------|------------------------|------------------------------
     // 01.00.00 19.08.2015  Siemens Industry Online Support
     //                      First released version
     // 01.00.01 02.01.2017  Siemens Industry Online Support
     //                      Upgrade: TIA Portal V14 Update 1
     // 01.00.02 17.08.2018  Siemens Industry Online Support
     //                      Upgrade: TIA V15 Update 2
     // 01.00.03 23.11.2018  Siemens Industry Online Support
     //                      Upgrade: TIA V15.1
     // 01.01.00 09.10.2019  Siemens Industry Presales Support
     //                      Renamed from "LGF_RandomInt" to "LGF_RandomRange_DInt"
     //                      change random datatype from int to dint
     //                      Regions, commens and costants are added
     // 03.00.00 23.04.2020  Siemens Industry Support
     //                      Set version to V3.0.0, harmonize the version of the whole library
     //=============================================================================
   END_REGION

   REGION Validation
     // Check if the maximal Value is less than the minimal value
     IF (#minValue > #maxValue) THEN
       #error := true;
       #status := #ERR_MAX_LESS_MIN;
       #subfunctionStatus := #SUB_STATUS_NO_ERROR;
       #LGF_RandomRange_Dint := #ZERO;
       RETURN;
     END_IF;

     // Read system time
     #tempTimeStatus := INT_TO_WORD(RD_SYS_T(#tempTime));

     // Check return variable for error
     IF (#tempTimeStatus <> #SUB_STATUS_NO_ERROR) THEN
       #error := true;
       #status := #ERR_RD_SYS_T;
       #subfunctionStatus := #tempTimeStatus;
       #LGF_RandomRange_Dint := #ZERO;
       RETURN;
     END_IF;
   END_REGION

   REGION Calculating random number
     // Converting to double word so individual bytes can be addressed
     #tempNanoSecondInDWord := UDINT_TO_DWORD(#tempTime.NANOSECOND);

     // Callculate a random-start-value depending on the time
     #tempRandomValue.%B3 := #tempNanoSecondInDWord.%B0;
     #tempRandomValue.%B2 := #tempNanoSecondInDWord.%B1;
     #tempRandomValue.%B1 := #tempNanoSecondInDWord.%B2;
     #tempRandomValue.%B0 := #tempNanoSecondInDWord.%B3;

     // Norm the calculated random number: 0.0 <= #tempNormReal <= 1.0
     #tempNormReal := UDINT_TO_REAL(DWORD_TO_UDINT(#tempRandomValue)) / UDINT_TO_REAL(#MAX_UDINT);

     // Scale the tempNormReal to be in the range of maxValue and minValue
     #LGF_RandomRange_Dint := REAL_TO_DINT((#tempNormReal * DINT_TO_REAL(#maxValue - #minValue) + DINT_TO_REAL(#minValue)));